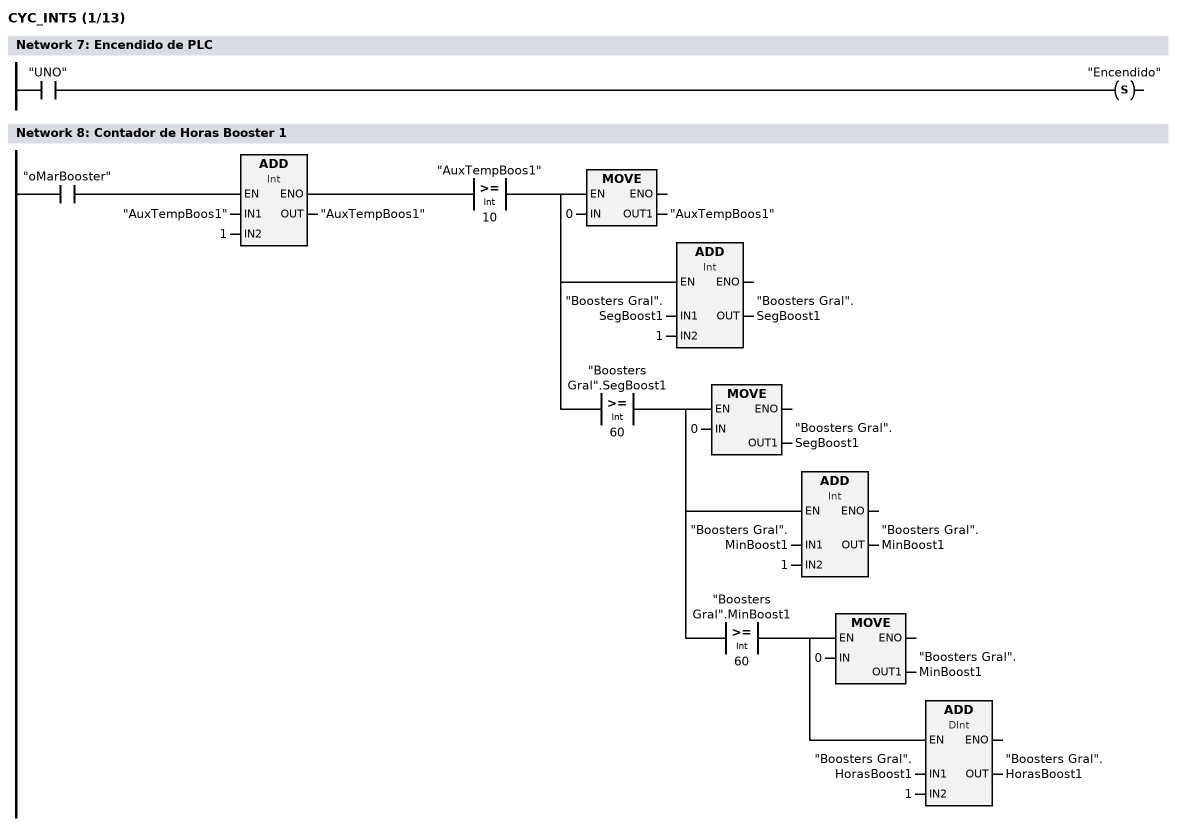
   RUNG wire#powerrail
      Contact( "UNO" )
      S_Coil( "Encendido" )
   END_RUNG
   // the same network as SCL:
   IF "UNO" THEN "Encendido" := TRUE; END_IF;
END_REGION

REGION Network 8: Contador de Horas Booster 1
   RUNG wire#powerrail
      Contact( "oMarBooster" )
      { S7_Templates := "SrcType := Int"; S7_GenerateENO := "TRUE" } Add(in1 := "AuxTempBoos1", in2 := 1, out => "AuxTempBoos1")
      { S7_Templates := "SrcType := Int" } GE_Contact(in1 := "AuxTempBoos1", in2 := 10)
      wire#w1
      { S7_GenerateENO := "TRUE" } Move(in := 0, out1 => "AuxTempBoos1")
   END_RUNG
   RUNG wire#w1
      { S7_Templates := "SrcType := Int"; S7_GenerateENO := "TRUE" } Add(in1 := "Boosters Gral".SegBoost1, in2 := 1, out => "Boosters Gral".SegBoost1)
   END_RUNG
   RUNG wire#w1
      { S7_Templates := "SrcType := Int" } GE_Contact(in1 := "Boosters Gral".SegBoost1, in2 := 60)
      wire#w2
      { S7_GenerateENO := "TRUE" } Move(in := 0, out1 => "Boosters Gral".SegBoost1)
   END_RUNG
   RUNG wire#w2
      { S7_Templates := "SrcType := Int"; S7_GenerateENO := "TRUE" } Add(in1 := "Boosters Gral".MinBoost1, in2 := 1, out => "Boosters Gral".MinBoost1)
   END_RUNG
   RUNG wire#w2
      { S7_Templates := "SrcType := Int" } GE_Contact(in1 := "Boosters Gral".MinBoost1, in2 := 60)
      wire#w3
      { S7_GenerateENO := "TRUE" } Move(in := 0, out1 => "Boosters Gral".MinBoost1)
   END_RUNG
   RUNG wire#w3
      { S7_Templates := "SrcType := DInt"; S7_GenerateENO := "TRUE" } Add(in1 := "Boosters Gral".HorasBoost1, in2 := 1, out => "Boosters Gral".HorasBoost1)
   END_RUNG
   // the same network as SCL:
   // ENO of a box is taken as its EN; it also drops when the box reports an error
   IF "oMarBooster" THEN "AuxTempBoos1" := "AuxTempBoos1" + 1; END_IF;
   #_w1 := "oMarBooster" AND ("AuxTempBoos1" >= 10);
   IF #_w1 THEN
       "AuxTempBoos1" := 0;
       "Boosters Gral".SegBoost1 := "Boosters Gral".SegBoost1 + 1;
   END_IF;
   #_w2 := #_w1 AND ("Boosters Gral".SegBoost1 >= 60);
   IF #_w2 THEN
       "Boosters Gral".SegBoost1 := 0;
       "Boosters Gral".MinBoost1 := "Boosters Gral".MinBoost1 + 1;
   END_IF;
   #_w3 := #_w2 AND ("Boosters Gral".MinBoost1 >= 60);
   IF #_w3 THEN
       "Boosters Gral".MinBoost1 := 0;
       "Boosters Gral".HorasBoost1 := "Boosters Gral".HorasBoost1 + 1;
   END_IF;
END_REGION

REGION Network 9: Contador de Horas Booster 2
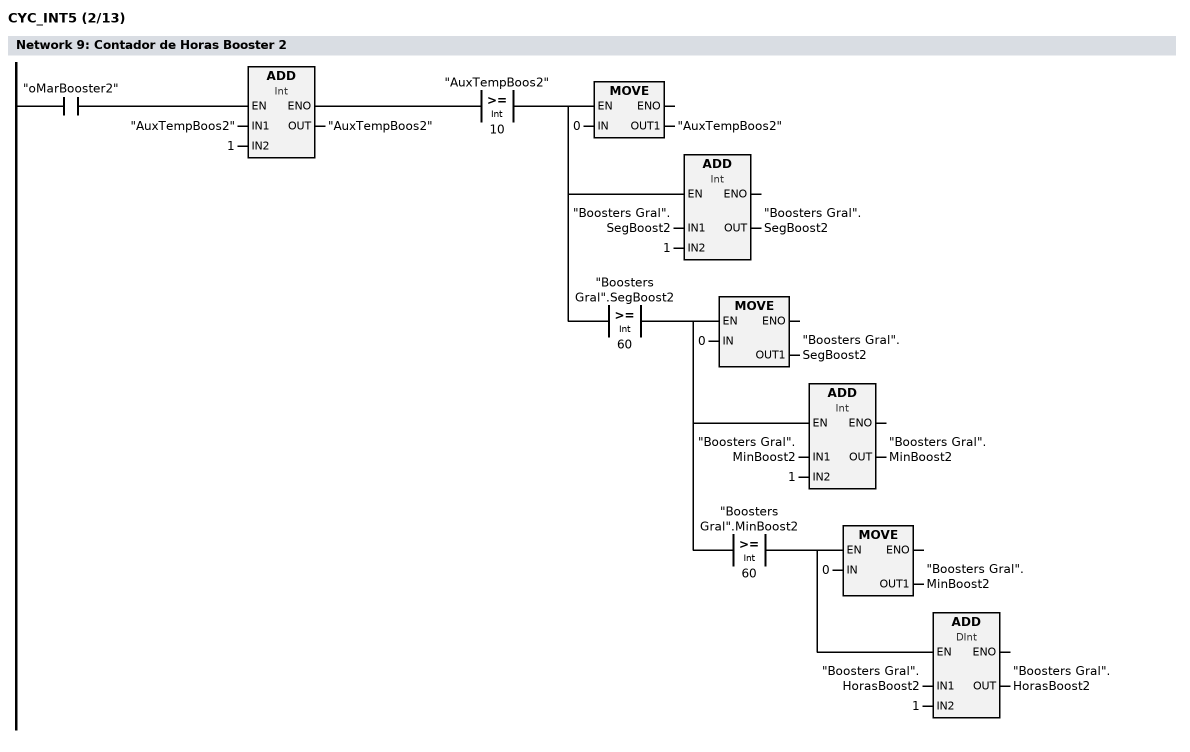
   RUNG wire#powerrail
      Contact( "oMarBooster2" )
      { S7_Templates := "SrcType := Int"; S7_GenerateENO := "TRUE" } Add(in1 := "AuxTempBoos2", in2 := 1, out => "AuxTempBoos2")
      { S7_Templates := "SrcType := Int" } GE_Contact(in1 := "AuxTempBoos2", in2 := 10)
      wire#w1
      { S7_GenerateENO := "TRUE" } Move(in := 0, out1 => "AuxTempBoos2")
   END_RUNG
   RUNG wire#w1
      { S7_Templates := "SrcType := Int"; S7_GenerateENO := "TRUE" } Add(in1 := "Boosters Gral".SegBoost2, in2 := 1, out => "Boosters Gral".SegBoost2)
   END_RUNG
   RUNG wire#w1
      { S7_Templates := "SrcType := Int" } GE_Contact(in1 := "Boosters Gral".SegBoost2, in2 := 60)
      wire#w2
      { S7_GenerateENO := "TRUE" } Move(in := 0, out1 => "Boosters Gral".SegBoost2)
   END_RUNG
   RUNG wire#w2
      { S7_Templates := "SrcType := Int"; S7_GenerateENO := "TRUE" } Add(in1 := "Boosters Gral".MinBoost2, in2 := 1, out => "Boosters Gral".MinBoost2)
   END_RUNG
   RUNG wire#w2
      { S7_Templates := "SrcType := Int" } GE_Contact(in1 := "Boosters Gral".MinBoost2, in2 := 60)
      wire#w3
      { S7_GenerateENO := "TRUE" } Move(in := 0, out1 => "Boosters Gral".MinBoost2)
   END_RUNG
   RUNG wire#w3
      { S7_Templates := "SrcType := DInt"; S7_GenerateENO := "TRUE" } Add(in1 := "Boosters Gral".HorasBoost2, in2 := 1, out => "Boosters Gral".HorasBoost2)
   END_RUNG
   // the same network as SCL:
   // ENO of a box is taken as its EN; it also drops when the box reports an error
   IF "oMarBooster2" THEN "AuxTempBoos2" := "AuxTempBoos2" + 1; END_IF;
   #_w1 := "oMarBooster2" AND ("AuxTempBoos2" >= 10);
   IF #_w1 THEN
       "AuxTempBoos2" := 0;
       "Boosters Gral".SegBoost2 := "Boosters Gral".SegBoost2 + 1;
   END_IF;
   #_w2 := #_w1 AND ("Boosters Gral".SegBoost2 >= 60);
   IF #_w2 THEN
       "Boosters Gral".SegBoost2 := 0;
       "Boosters Gral".MinBoost2 := "Boosters Gral".MinBoost2 + 1;
   END_IF;
   #_w3 := #_w2 AND ("Boosters Gral".MinBoost2 >= 60);
   IF #_w3 THEN
       "Boosters Gral".MinBoost2 := 0;
       "Boosters Gral".HorasBoost2 := "Boosters Gral".HorasBoost2 + 1;
   END_IF;
END_REGION

REGION Network 10: Horas de marcha MS050 / Contador de Horas Booster 1
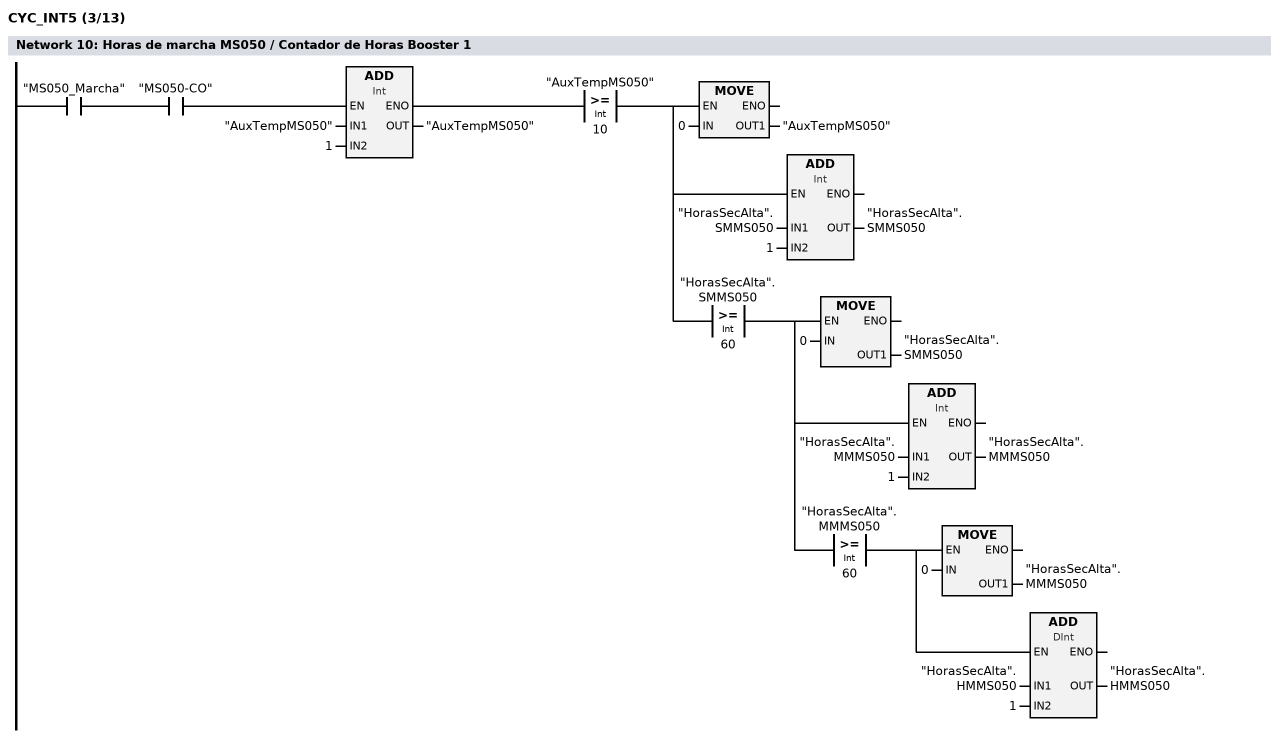
   RUNG wire#powerrail
      Contact( "MS050_Marcha" )
      Contact( "MS050-CO" )
      { S7_Templates := "SrcType := Int"; S7_GenerateENO := "TRUE" } Add(in1 := "AuxTempMS050", in2 := 1, out => "AuxTempMS050")
      { S7_Templates := "SrcType := Int" } GE_Contact(in1 := "AuxTempMS050", in2 := 10)
      wire#w1
      { S7_GenerateENO := "TRUE" } Move(in := 0, out1 => "AuxTempMS050")
   END_RUNG
   RUNG wire#w1
      { S7_Templates := "SrcType := Int"; S7_GenerateENO := "TRUE" } Add(in1 := "HorasSecAlta".SMMS050, in2 := 1, out => "HorasSecAlta".SMMS050)
   END_RUNG
   RUNG wire#w1
      { S7_Templates := "SrcType := Int" } GE_Contact(in1 := "HorasSecAlta".SMMS050, in2 := 60)
      wire#w2
      { S7_GenerateENO := "TRUE" } Move(in := 0, out1 => "HorasSecAlta".SMMS050)
   END_RUNG
   RUNG wire#w2
      { S7_Templates := "SrcType := Int"; S7_GenerateENO := "TRUE" } Add(in1 := "HorasSecAlta".MMMS050, in2 := 1, out => "HorasSecAlta".MMMS050)
   END_RUNG
   RUNG wire#w2
      { S7_Templates := "SrcType := Int" } GE_Contact(in1 := "HorasSecAlta".MMMS050, in2 := 60)
      wire#w3
      { S7_GenerateENO := "TRUE" } Move(in := 0, out1 => "HorasSecAlta".MMMS050)
   END_RUNG
   RUNG wire#w3
      { S7_Templates := "SrcType := DInt"; S7_GenerateENO := "TRUE" } Add(in1 := "HorasSecAlta".HMMS050, in2 := 1, out => "HorasSecAlta".HMMS050)
   END_RUNG
   // the same network as SCL:
   // ENO of a box is taken as its EN; it also drops when the box reports an error
   #_w1 := "MS050_Marcha" AND "MS050-CO";
   IF #_w1 THEN "AuxTempMS050" := "AuxTempMS050" + 1; END_IF;
   #_w2 := #_w1 AND ("AuxTempMS050" >= 10);
   IF #_w2 THEN
       "AuxTempMS050" := 0;
       "HorasSecAlta".SMMS050 := "HorasSecAlta".SMMS050 + 1;
   END_IF;
   #_w3 := #_w2 AND ("HorasSecAlta".SMMS050 >= 60);
   IF #_w3 THEN
       "HorasSecAlta".SMMS050 := 0;
       "HorasSecAlta".MMMS050 := "HorasSecAlta".MMMS050 + 1;
   END_IF;
   #_w4 := #_w3 AND ("HorasSecAlta".MMMS050 >= 60);
   IF #_w4 THEN
       "HorasSecAlta".MMMS050 := 0;
       "HorasSecAlta".HMMS050 := "HorasSecAlta".HMMS050 + 1;
   END_IF;
END_REGION

REGION Network 11: Horas de marcha MS051 / Contador de Horas Booster 1
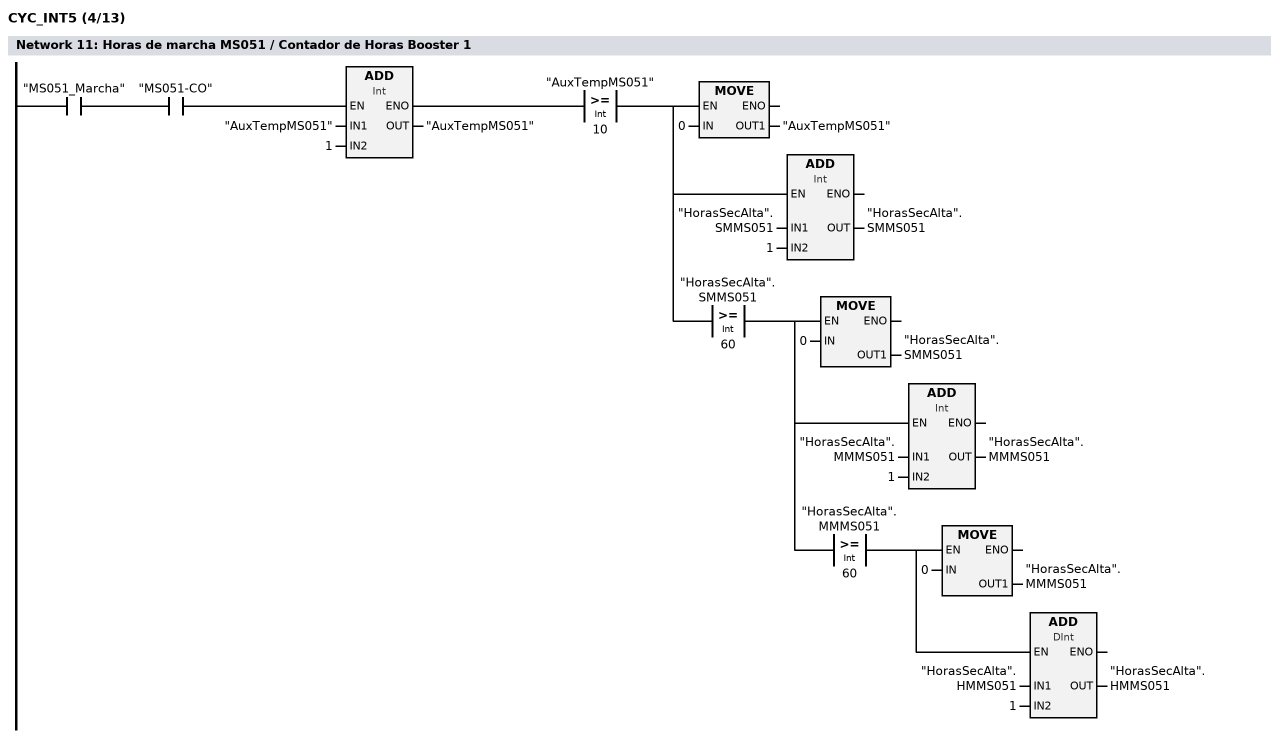
   RUNG wire#powerrail
      Contact( "MS051_Marcha" )
      Contact( "MS051-CO" )
      { S7_Templates := "SrcType := Int"; S7_GenerateENO := "TRUE" } Add(in1 := "AuxTempMS051", in2 := 1, out => "AuxTempMS051")
      { S7_Templates := "SrcType := Int" } GE_Contact(in1 := "AuxTempMS051", in2 := 10)
      wire#w1
      { S7_GenerateENO := "TRUE" } Move(in := 0, out1 => "AuxTempMS051")
   END_RUNG
   RUNG wire#w1
      { S7_Templates := "SrcType := Int"; S7_GenerateENO := "TRUE" } Add(in1 := "HorasSecAlta".SMMS051, in2 := 1, out => "HorasSecAlta".SMMS051)
   END_RUNG
   RUNG wire#w1
      { S7_Templates := "SrcType := Int" } GE_Contact(in1 := "HorasSecAlta".SMMS051, in2 := 60)
      wire#w2
      { S7_GenerateENO := "TRUE" } Move(in := 0, out1 => "HorasSecAlta".SMMS051)
   END_RUNG
   RUNG wire#w2
      { S7_Templates := "SrcType := Int"; S7_GenerateENO := "TRUE" } Add(in1 := "HorasSecAlta".MMMS051, in2 := 1, out => "HorasSecAlta".MMMS051)
   END_RUNG
   RUNG wire#w2
      { S7_Templates := "SrcType := Int" } GE_Contact(in1 := "HorasSecAlta".MMMS051, in2 := 60)
      wire#w3
      { S7_GenerateENO := "TRUE" } Move(in := 0, out1 => "HorasSecAlta".MMMS051)
   END_RUNG
   RUNG wire#w3
      { S7_Templates := "SrcType := DInt"; S7_GenerateENO := "TRUE" } Add(in1 := "HorasSecAlta".HMMS051, in2 := 1, out => "HorasSecAlta".HMMS051)
   END_RUNG
   // the same network as SCL:
   // ENO of a box is taken as its EN; it also drops when the box reports an error
   #_w1 := "MS051_Marcha" AND "MS051-CO";
   IF #_w1 THEN "AuxTempMS051" := "AuxTempMS051" + 1; END_IF;
   #_w2 := #_w1 AND ("AuxTempMS051" >= 10);
   IF #_w2 THEN
       "AuxTempMS051" := 0;
       "HorasSecAlta".SMMS051 := "HorasSecAlta".SMMS051 + 1;
   END_IF;
   #_w3 := #_w2 AND ("HorasSecAlta".SMMS051 >= 60);
   IF #_w3 THEN
       "HorasSecAlta".SMMS051 := 0;
       "HorasSecAlta".MMMS051 := "HorasSecAlta".MMMS051 + 1;
   END_IF;
   #_w4 := #_w3 AND ("HorasSecAlta".MMMS051 >= 60);
   IF #_w4 THEN
       "HorasSecAlta".MMMS051 := 0;
       "HorasSecAlta".HMMS051 := "HorasSecAlta".HMMS051 + 1;
   END_IF;
END_REGION

REGION Network 12: Horas de marcha MS052 / Contador de Horas Booster 1
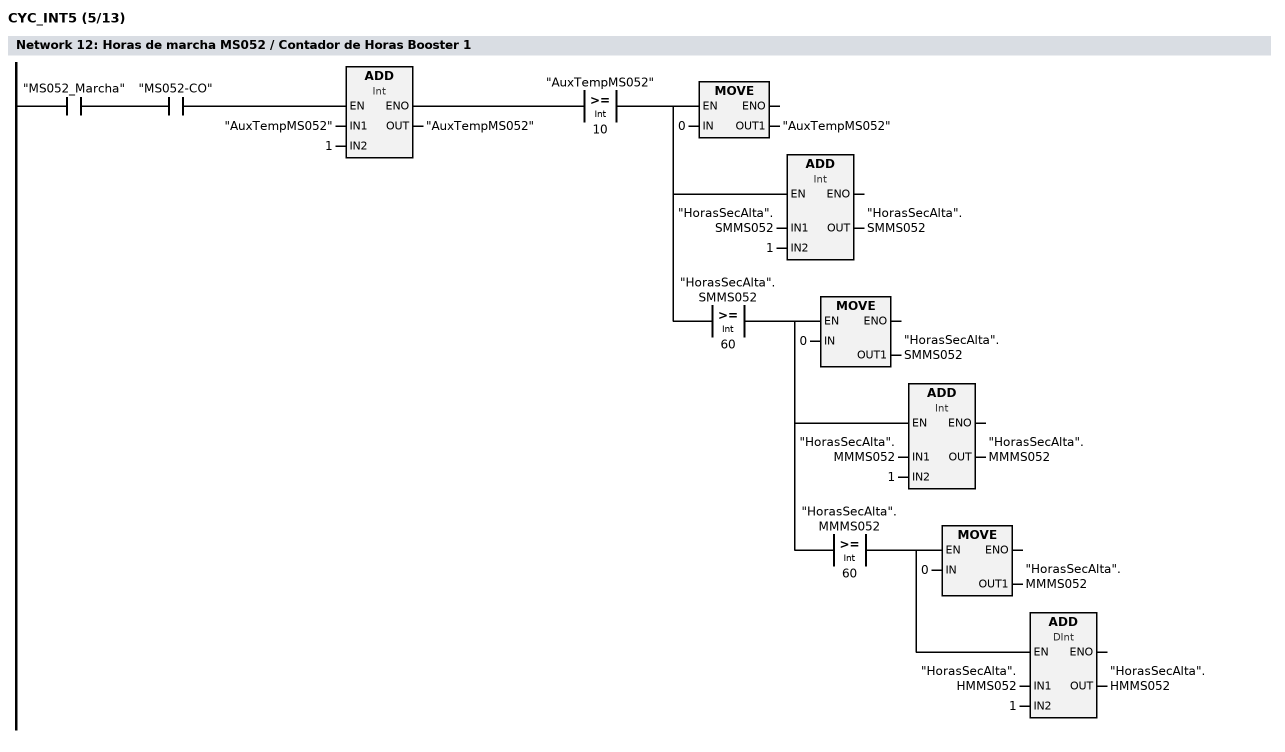
   RUNG wire#powerrail
      Contact( "MS052_Marcha" )
      Contact( "MS052-CO" )
      { S7_Templates := "SrcType := Int"; S7_GenerateENO := "TRUE" } Add(in1 := "AuxTempMS052", in2 := 1, out => "AuxTempMS052")
      { S7_Templates := "SrcType := Int" } GE_Contact(in1 := "AuxTempMS052", in2 := 10)
      wire#w1
      { S7_GenerateENO := "TRUE" } Move(in := 0, out1 => "AuxTempMS052")
   END_RUNG
   RUNG wire#w1
      { S7_Templates := "SrcType := Int"; S7_GenerateENO := "TRUE" } Add(in1 := "HorasSecAlta".SMMS052, in2 := 1, out => "HorasSecAlta".SMMS052)
   END_RUNG
   RUNG wire#w1
      { S7_Templates := "SrcType := Int" } GE_Contact(in1 := "HorasSecAlta".SMMS052, in2 := 60)
      wire#w2
      { S7_GenerateENO := "TRUE" } Move(in := 0, out1 => "HorasSecAlta".SMMS052)
   END_RUNG
   RUNG wire#w2
      { S7_Templates := "SrcType := Int"; S7_GenerateENO := "TRUE" } Add(in1 := "HorasSecAlta".MMMS052, in2 := 1, out => "HorasSecAlta".MMMS052)
   END_RUNG
   RUNG wire#w2
      { S7_Templates := "SrcType := Int" } GE_Contact(in1 := "HorasSecAlta".MMMS052, in2 := 60)
      wire#w3
      { S7_GenerateENO := "TRUE" } Move(in := 0, out1 => "HorasSecAlta".MMMS052)
   END_RUNG
   RUNG wire#w3
      { S7_Templates := "SrcType := DInt"; S7_GenerateENO := "TRUE" } Add(in1 := "HorasSecAlta".HMMS052, in2 := 1, out => "HorasSecAlta".HMMS052)
   END_RUNG
   // the same network as SCL:
   // ENO of a box is taken as its EN; it also drops when the box reports an error
   #_w1 := "MS052_Marcha" AND "MS052-CO";
   IF #_w1 THEN "AuxTempMS052" := "AuxTempMS052" + 1; END_IF;
   #_w2 := #_w1 AND ("AuxTempMS052" >= 10);
   IF #_w2 THEN
       "AuxTempMS052" := 0;
       "HorasSecAlta".SMMS052 := "HorasSecAlta".SMMS052 + 1;
   END_IF;
   #_w3 := #_w2 AND ("HorasSecAlta".SMMS052 >= 60);
   IF #_w3 THEN
       "HorasSecAlta".SMMS052 := 0;
       "HorasSecAlta".MMMS052 := "HorasSecAlta".MMMS052 + 1;
   END_IF;
   #_w4 := #_w3 AND ("HorasSecAlta".MMMS052 >= 60);
   IF #_w4 THEN
       "HorasSecAlta".MMMS052 := 0;
       "HorasSecAlta".HMMS052 := "HorasSecAlta".HMMS052 + 1;
   END_IF;
END_REGION

REGION Network 13: Horas de marcha MS053 / Contador de Horas Booster 1
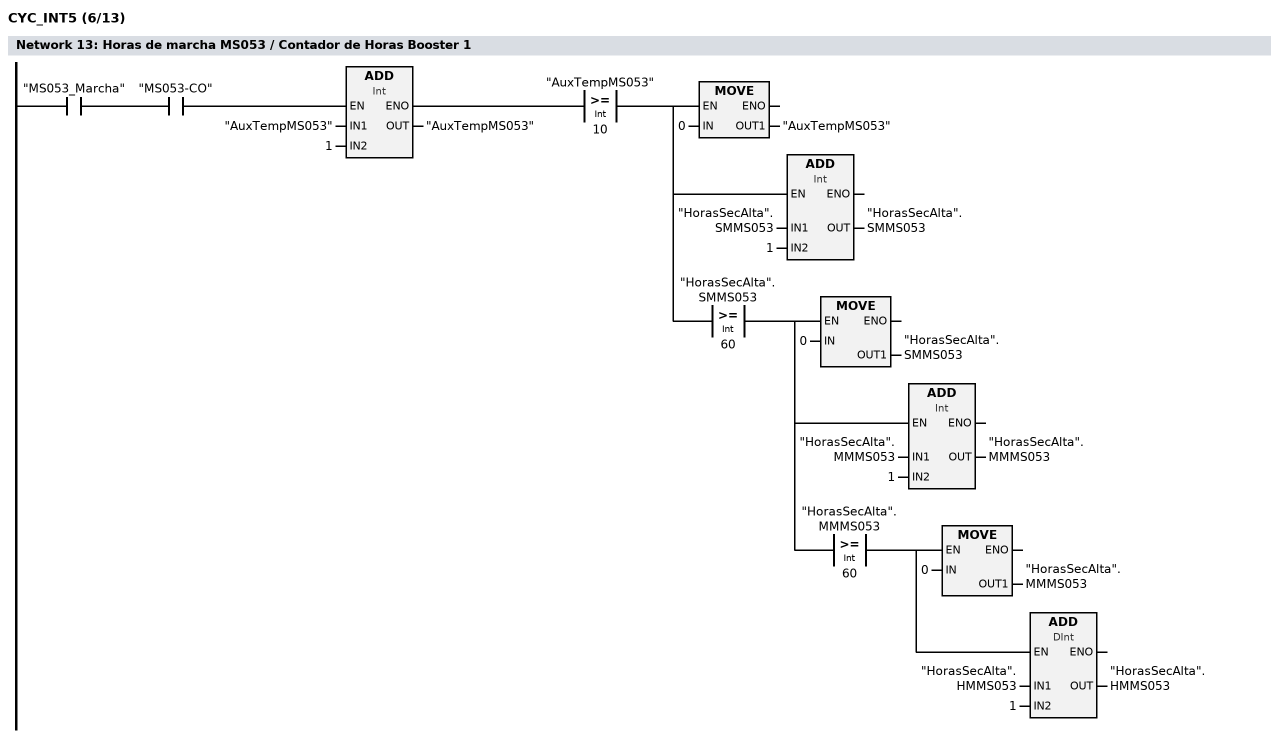
   RUNG wire#powerrail
      Contact( "MS053_Marcha" )
      Contact( "MS053-CO" )
      { S7_Templates := "SrcType := Int"; S7_GenerateENO := "TRUE" } Add(in1 := "AuxTempMS053", in2 := 1, out => "AuxTempMS053")
      { S7_Templates := "SrcType := Int" } GE_Contact(in1 := "AuxTempMS053", in2 := 10)
      wire#w1
      { S7_GenerateENO := "TRUE" } Move(in := 0, out1 => "AuxTempMS053")
   END_RUNG
   RUNG wire#w1
      { S7_Templates := "SrcType := Int"; S7_GenerateENO := "TRUE" } Add(in1 := "HorasSecAlta".SMMS053, in2 := 1, out => "HorasSecAlta".SMMS053)
   END_RUNG
   RUNG wire#w1
      { S7_Templates := "SrcType := Int" } GE_Contact(in1 := "HorasSecAlta".SMMS053, in2 := 60)
      wire#w2
      { S7_GenerateENO := "TRUE" } Move(in := 0, out1 => "HorasSecAlta".SMMS053)
   END_RUNG
   RUNG wire#w2
      { S7_Templates := "SrcType := Int"; S7_GenerateENO := "TRUE" } Add(in1 := "HorasSecAlta".MMMS053, in2 := 1, out => "HorasSecAlta".MMMS053)
   END_RUNG
   RUNG wire#w2
      { S7_Templates := "SrcType := Int" } GE_Contact(in1 := "HorasSecAlta".MMMS053, in2 := 60)
      wire#w3
      { S7_GenerateENO := "TRUE" } Move(in := 0, out1 => "HorasSecAlta".MMMS053)
   END_RUNG
   RUNG wire#w3
      { S7_Templates := "SrcType := DInt"; S7_GenerateENO := "TRUE" } Add(in1 := "HorasSecAlta".HMMS053, in2 := 1, out => "HorasSecAlta".HMMS053)
   END_RUNG
   // the same network as SCL:
   // ENO of a box is taken as its EN; it also drops when the box reports an error
   #_w1 := "MS053_Marcha" AND "MS053-CO";
   IF #_w1 THEN "AuxTempMS053" := "AuxTempMS053" + 1; END_IF;
   #_w2 := #_w1 AND ("AuxTempMS053" >= 10);
   IF #_w2 THEN
       "AuxTempMS053" := 0;
       "HorasSecAlta".SMMS053 := "HorasSecAlta".SMMS053 + 1;
   END_IF;
   #_w3 := #_w2 AND ("HorasSecAlta".SMMS053 >= 60);
   IF #_w3 THEN
       "HorasSecAlta".SMMS053 := 0;
       "HorasSecAlta".MMMS053 := "HorasSecAlta".MMMS053 + 1;
   END_IF;
   #_w4 := #_w3 AND ("HorasSecAlta".MMMS053 >= 60);
   IF #_w4 THEN
       "HorasSecAlta".MMMS053 := 0;
       "HorasSecAlta".HMMS053 := "HorasSecAlta".HMMS053 + 1;
   END_IF;
END_REGION

REGION Network 14: Horas de marcha MS054 / Contador de Horas Booster 1
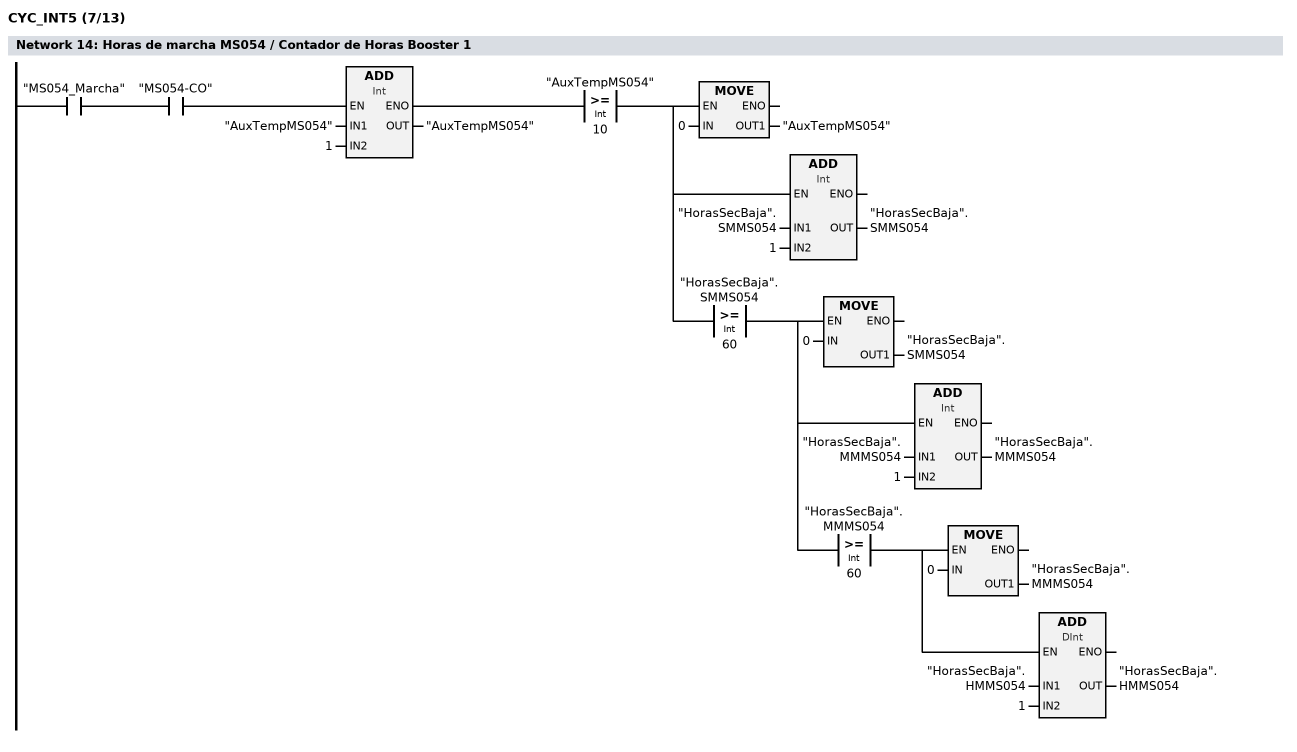
   RUNG wire#powerrail
      Contact( "MS054_Marcha" )
      Contact( "MS054-CO" )
      { S7_Templates := "SrcType := Int"; S7_GenerateENO := "TRUE" } Add(in1 := "AuxTempMS054", in2 := 1, out => "AuxTempMS054")
      { S7_Templates := "SrcType := Int" } GE_Contact(in1 := "AuxTempMS054", in2 := 10)
      wire#w1
      { S7_GenerateENO := "TRUE" } Move(in := 0, out1 => "AuxTempMS054")
   END_RUNG
   RUNG wire#w1
      { S7_Templates := "SrcType := Int"; S7_GenerateENO := "TRUE" } Add(in1 := "HorasSecBaja".SMMS054, in2 := 1, out => "HorasSecBaja".SMMS054)
   END_RUNG
   RUNG wire#w1
      { S7_Templates := "SrcType := Int" } GE_Contact(in1 := "HorasSecBaja".SMMS054, in2 := 60)
      wire#w2
      { S7_GenerateENO := "TRUE" } Move(in := 0, out1 => "HorasSecBaja".SMMS054)
   END_RUNG
   RUNG wire#w2
      { S7_Templates := "SrcType := Int"; S7_GenerateENO := "TRUE" } Add(in1 := "HorasSecBaja".MMMS054, in2 := 1, out => "HorasSecBaja".MMMS054)
   END_RUNG
   RUNG wire#w2
      { S7_Templates := "SrcType := Int" } GE_Contact(in1 := "HorasSecBaja".MMMS054, in2 := 60)
      wire#w3
      { S7_GenerateENO := "TRUE" } Move(in := 0, out1 => "HorasSecBaja".MMMS054)
   END_RUNG
   RUNG wire#w3
      { S7_Templates := "SrcType := DInt"; S7_GenerateENO := "TRUE" } Add(in1 := "HorasSecBaja".HMMS054, in2 := 1, out => "HorasSecBaja".HMMS054)
   END_RUNG
   // the same network as SCL:
   // ENO of a box is taken as its EN; it also drops when the box reports an error
   #_w1 := "MS054_Marcha" AND "MS054-CO";
   IF #_w1 THEN "AuxTempMS054" := "AuxTempMS054" + 1; END_IF;
   #_w2 := #_w1 AND ("AuxTempMS054" >= 10);
   IF #_w2 THEN
       "AuxTempMS054" := 0;
       "HorasSecBaja".SMMS054 := "HorasSecBaja".SMMS054 + 1;
   END_IF;
   #_w3 := #_w2 AND ("HorasSecBaja".SMMS054 >= 60);
   IF #_w3 THEN
       "HorasSecBaja".SMMS054 := 0;
       "HorasSecBaja".MMMS054 := "HorasSecBaja".MMMS054 + 1;
   END_IF;
   #_w4 := #_w3 AND ("HorasSecBaja".MMMS054 >= 60);
   IF #_w4 THEN
       "HorasSecBaja".MMMS054 := 0;
       "HorasSecBaja".HMMS054 := "HorasSecBaja".HMMS054 + 1;
   END_IF;
END_REGION

REGION Network 15: Horas de marcha MS055 / Contador de Horas Booster 1
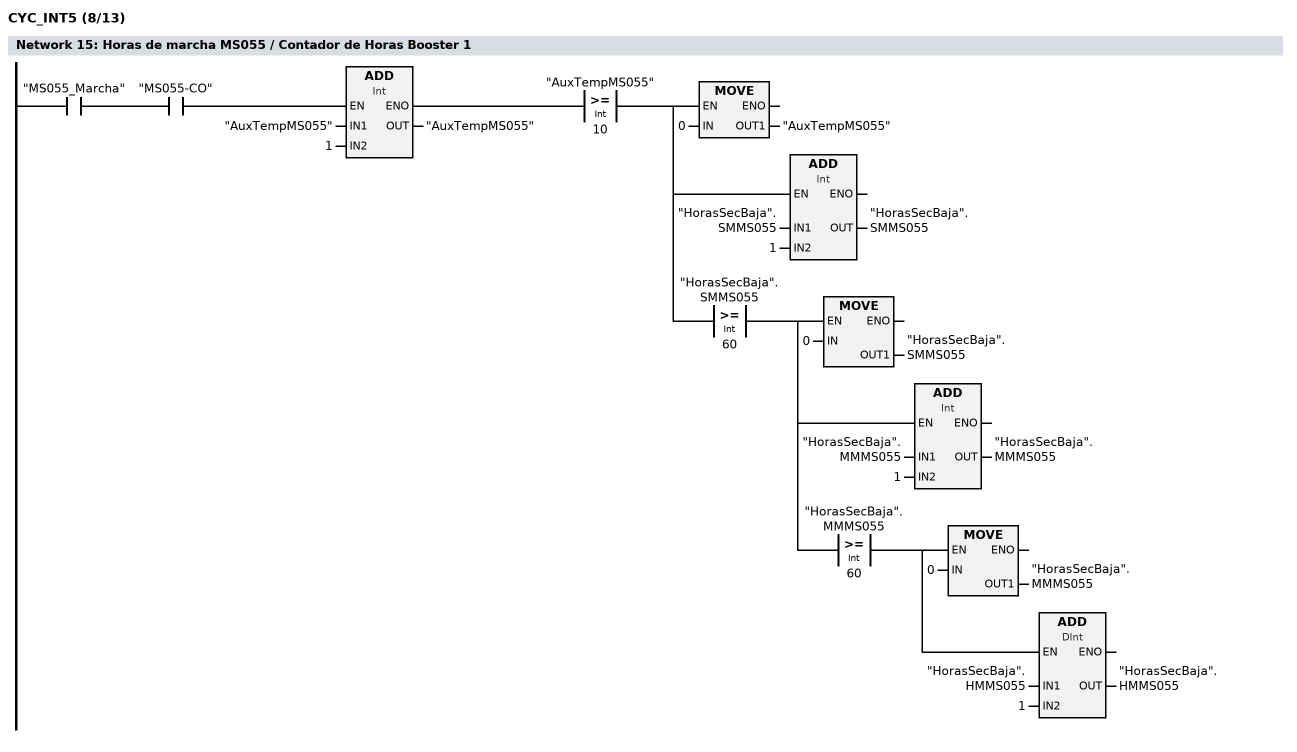
   RUNG wire#powerrail
      Contact( "MS055_Marcha" )
      Contact( "MS055-CO" )
      { S7_Templates := "SrcType := Int"; S7_GenerateENO := "TRUE" } Add(in1 := "AuxTempMS055", in2 := 1, out => "AuxTempMS055")
      { S7_Templates := "SrcType := Int" } GE_Contact(in1 := "AuxTempMS055", in2 := 10)
      wire#w1
      { S7_GenerateENO := "TRUE" } Move(in := 0, out1 => "AuxTempMS055")
   END_RUNG
   RUNG wire#w1
      { S7_Templates := "SrcType := Int"; S7_GenerateENO := "TRUE" } Add(in1 := "HorasSecBaja".SMMS055, in2 := 1, out => "HorasSecBaja".SMMS055)
   END_RUNG
   RUNG wire#w1
      { S7_Templates := "SrcType := Int" } GE_Contact(in1 := "HorasSecBaja".SMMS055, in2 := 60)
      wire#w2
      { S7_GenerateENO := "TRUE" } Move(in := 0, out1 => "HorasSecBaja".SMMS055)
   END_RUNG
   RUNG wire#w2
      { S7_Templates := "SrcType := Int"; S7_GenerateENO := "TRUE" } Add(in1 := "HorasSecBaja".MMMS055, in2 := 1, out => "HorasSecBaja".MMMS055)
   END_RUNG
   RUNG wire#w2
      { S7_Templates := "SrcType := Int" } GE_Contact(in1 := "HorasSecBaja".MMMS055, in2 := 60)
      wire#w3
      { S7_GenerateENO := "TRUE" } Move(in := 0, out1 => "HorasSecBaja".MMMS055)
   END_RUNG
   RUNG wire#w3
      { S7_Templates := "SrcType := DInt"; S7_GenerateENO := "TRUE" } Add(in1 := "HorasSecBaja".HMMS055, in2 := 1, out => "HorasSecBaja".HMMS055)
   END_RUNG
   // the same network as SCL:
   // ENO of a box is taken as its EN; it also drops when the box reports an error
   #_w1 := "MS055_Marcha" AND "MS055-CO";
   IF #_w1 THEN "AuxTempMS055" := "AuxTempMS055" + 1; END_IF;
   #_w2 := #_w1 AND ("AuxTempMS055" >= 10);
   IF #_w2 THEN
       "AuxTempMS055" := 0;
       "HorasSecBaja".SMMS055 := "HorasSecBaja".SMMS055 + 1;
   END_IF;
   #_w3 := #_w2 AND ("HorasSecBaja".SMMS055 >= 60);
   IF #_w3 THEN
       "HorasSecBaja".SMMS055 := 0;
       "HorasSecBaja".MMMS055 := "HorasSecBaja".MMMS055 + 1;
   END_IF;
   #_w4 := #_w3 AND ("HorasSecBaja".MMMS055 >= 60);
   IF #_w4 THEN
       "HorasSecBaja".MMMS055 := 0;
       "HorasSecBaja".HMMS055 := "HorasSecBaja".HMMS055 + 1;
   END_IF;
END_REGION

REGION Network 16: Horas de marcha MC060 / Contador de Horas Booster 1